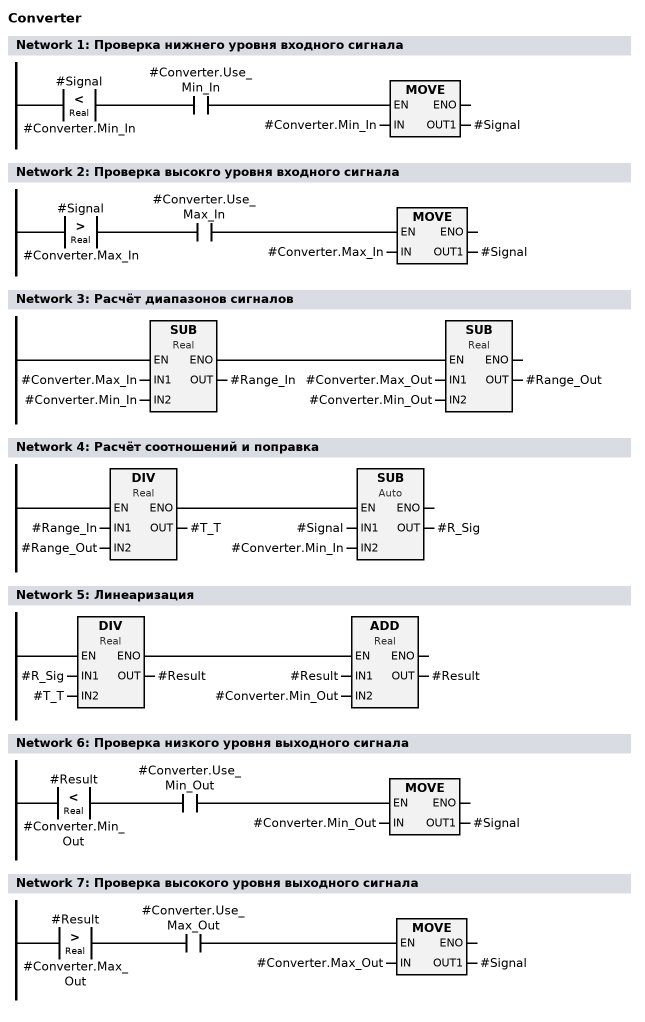
   RUNG wire#powerrail
      { S7_Templates := "SrcType := Real" } LT_Contact(in1 := #Signal, in2 := #Converter.Min_In)
      Contact( #Converter.Use_Min_In )
      Move(in := #Converter.Min_In, out1 => #Signal)
   END_RUNG
   // the same network as SCL:
   IF (#Signal < #Converter.Min_In) AND #Converter.Use_Min_In THEN #Signal := #Converter.Min_In; END_IF;
END_REGION

REGION Network 2: Проверка высокго уровня входного сигнала
   RUNG wire#powerrail
      { S7_Templates := "SrcType := Real" } GT_Contact(in1 := #Signal, in2 := #Converter.Max_In)
      Contact( #Converter.Use_Max_In )
      Move(in := #Converter.Max_In, out1 => #Signal)
   END_RUNG
   // the same network as SCL:
   IF (#Signal > #Converter.Max_In) AND #Converter.Use_Max_In THEN #Signal := #Converter.Max_In; END_IF;
END_REGION

REGION Network 3: Расчёт диапазонов сигналов
   RUNG wire#powerrail
      { S7_Templates := "SrcType := Real"; S7_GenerateENO := "TRUE" } Sub(in1 := #Converter.Max_In, in2 := #Converter.Min_In, out => #Range_In)
      { S7_Templates := "SrcType := Real"; S7_GenerateENO := "TRUE" } Sub(in1 := #Converter.Max_Out, in2 := #Converter.Min_Out, out => #Range_Out)
   END_RUNG
   // the same network as SCL:
   // ENO of a box is taken as its EN; it also drops when the box reports an error
   #Range_In := #Converter.Max_In - #Converter.Min_In;
   #Range_Out := #Converter.Max_Out - #Converter.Min_Out;
END_REGION

REGION Network 4: Расчёт соотношений и поправка
   RUNG wire#powerrail
      { S7_Templates := "SrcType := Real"; S7_GenerateENO := "TRUE" } Div(in1 := #Range_In, in2 := #Range_Out, out => #T_T)
      Sub(in1 := #Signal, in2 := #Converter.Min_In, out => #R_Sig)
   END_RUNG
   // the same network as SCL:
   // ENO of a box is taken as its EN; it also drops when the box reports an error
   #T_T := #Range_In / #Range_Out;
   #R_Sig := #Signal - #Converter.Min_In;
END_REGION

REGION Network 5: Линеаризация
   RUNG wire#powerrail
      { S7_Templates := "SrcType := Real"; S7_GenerateENO := "TRUE" } Div(in1 := #R_Sig, in2 := #T_T, out => #Result)
      { S7_Templates := "SrcType := Real"; S7_GenerateENO := "TRUE" } Add(in1 := #Result, in2 := #Converter.Min_Out, out => #Result)
   END_RUNG
   // the same network as SCL:
   // ENO of a box is taken as its EN; it also drops when the box reports an error
   #Result := #R_Sig / #T_T;
   #Result := #Result + #Converter.Min_Out;
END_REGION

REGION Network 6: Проверка низкого уровня выходного сигнала
   RUNG wire#powerrail
      { S7_Templates := "SrcType := Real" } LT_Contact(in1 := #Result, in2 := #Converter.Min_Out)
      Contact( #Converter.Use_Min_Out )
      Move(in := #Converter.Min_Out, out1 => #Signal)
   END_RUNG
   // the same network as SCL:
   IF (#Result < #Converter.Min_Out) AND #Converter.Use_Min_Out THEN #Signal := #Converter.Min_Out; END_IF;
END_REGION

REGION Network 7: Проверка высокого уровня выходного сигнала
   RUNG wire#powerrail
      { S7_Templates := "SrcType := Real" } GT_Contact(in1 := #Result, in2 := #Converter.Max_Out)
      Contact( #Converter.Use_Max_Out )
      Move(in := #Converter.Max_Out, out1 => #Signal)
   END_RUNG
   // the same network as SCL:
   IF (#Result > #Converter.Max_Out) AND #Converter.Use_Max_Out THEN #Signal := #Converter.Max_Out; END_IF;
END_REGION
END_FUNCTION

FUNCTION "INV" : Void   // FC111, LAD
{ S7_Optimized_Access := 'TRUE' }
VERSION : 0.1
   VAR_INPUT
      S : Bool;   // Сигнал
      I : Bool;   // Инверсия
   END_VAR
   VAR_IN_OUT
      R : Bool;   // Результат
   END_VAR
BEGIN

REGION Network 1: Инверсия сигнала
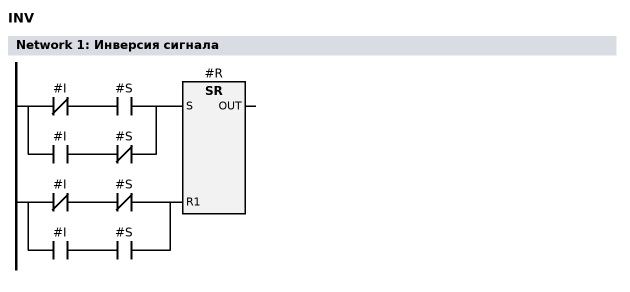
   RUNG wire#powerrail
      I_Contact( #I )
      Contact( #S )
      wire#w1
      S_SR(operand := #R, r1 := wire#w2)
   END_RUNG
   RUNG wire#powerrail
      Contact( #I )
      I_Contact( #S )
   END_RUNG wire#w1
   RUNG wire#powerrail
      I_Contact( #I )
      I_Contact( #S )
   END_RUNG wire#w2
   RUNG wire#powerrail
      Contact( #I )
      Contact( #S )
   END_RUNG wire#w2
   // the same network as SCL:
   IF (NOT #I AND #S) OR (#I AND NOT #S) THEN
       #R := TRUE;   // SR flip-flop
   END_IF;
   IF (NOT #I AND NOT #S) OR (#I AND #S) THEN #R := FALSE; END_IF;
END_REGION
END_FUNCTION

FUNCTION "Mode" : Void   // FC150, LAD
{ S7_Optimized_Access := 'FALSE' }
VERSION : 0.1
   VAR_INPUT
      CMD : Struct   // Основные команды
         Hand : Bool;   // 0 - авто, 1 - ручной / 0 - Авто, 1 - Ручной
         Start_A : Bool;   // Автозапуск / Запуск в авторежиме
         Start_M : Bool;   // Ручной - вперёд / Запуск в ручном режиме
         Force : Bool;   // Принудительный
         Lock : Bool;   // Блокировать / Блокировка
         Local : Bool;   // Локальный
         Service : Bool;   // Сервис
         Safety : Bool;   // Безопасность
         Alarm : Bool;   // Есть авария / Авария
         Reset : Bool;   // Сброс аварий
         Sim : Bool;   // Режим симуляции
      END_STRUCT;
      All_Block : Bool;   // Аварийная блокировка
   END_VAR
   VAR_OUTPUT
      Mode : Int;   // Режим работы
   END_VAR
BEGIN

REGION Network 1: Автоматический режим
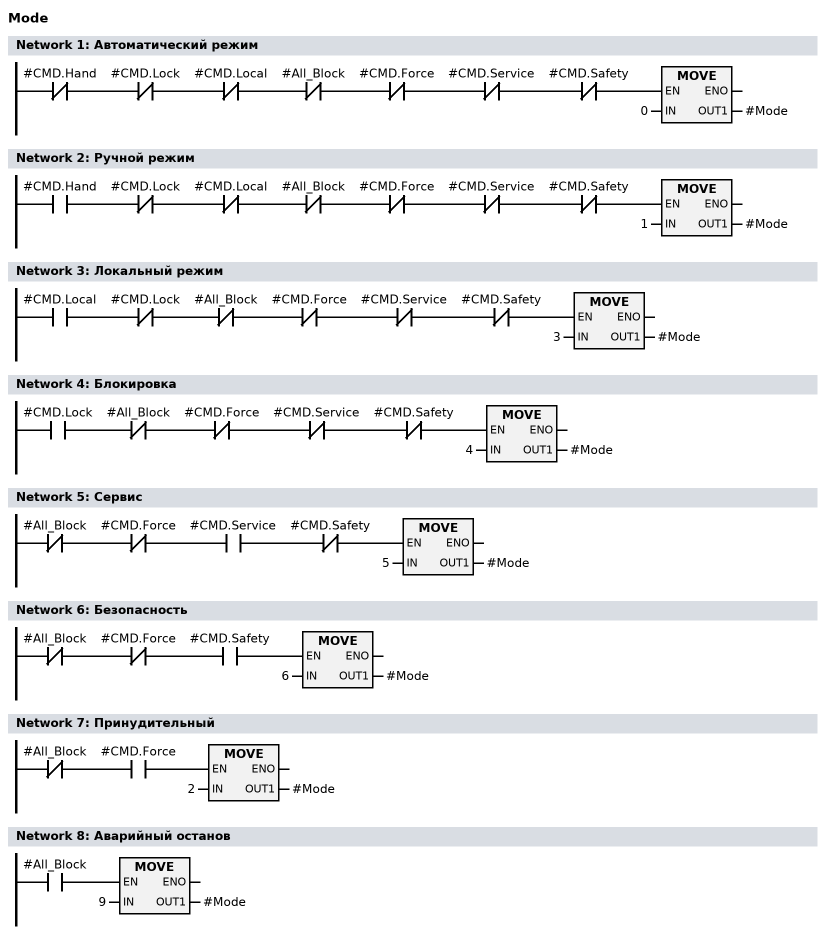
   RUNG wire#powerrail
      I_Contact( #CMD.Hand )
      I_Contact( #CMD.Lock )
      I_Contact( #CMD.Local )
      I_Contact( #All_Block )
      I_Contact( #CMD.Force )
      I_Contact( #CMD.Service )
      I_Contact( #CMD.Safety )
      { S7_GenerateENO := "TRUE" } Move(in := 0, out1 => #Mode)
   END_RUNG
   // the same network as SCL:
   IF NOT #CMD.Hand AND NOT #CMD.Lock AND NOT #CMD.Local AND NOT #All_Block AND NOT #CMD.Force AND NOT #CMD.Service AND NOT #CMD.Safety THEN
       #Mode := 0;
   END_IF;
END_REGION

REGION Network 2: Ручной режим
   RUNG wire#powerrail
      Contact( #CMD.Hand )
      I_Contact( #CMD.Lock )
      I_Contact( #CMD.Local )
      I_Contact( #All_Block )
      I_Contact( #CMD.Force )
      I_Contact( #CMD.Service )
      I_Contact( #CMD.Safety )
      { S7_GenerateENO := "TRUE" } Move(in := 1, out1 => #Mode)
   END_RUNG
   // the same network as SCL:
   IF #CMD.Hand AND NOT #CMD.Lock AND NOT #CMD.Local AND NOT #All_Block AND NOT #CMD.Force AND NOT #CMD.Service AND NOT #CMD.Safety THEN
       #Mode := 1;
   END_IF;
END_REGION

REGION Network 3: Локальный режим
   RUNG wire#powerrail
      Contact( #CMD.Local )
      I_Contact( #CMD.Lock )
      I_Contact( #All_Block )
      I_Contact( #CMD.Force )
      I_Contact( #CMD.Service )
      I_Contact( #CMD.Safety )
      { S7_GenerateENO := "TRUE" } Move(in := 3, out1 => #Mode)
   END_RUNG
   // the same network as SCL:
   IF #CMD.Local AND NOT #CMD.Lock AND NOT #All_Block AND NOT #CMD.Force AND NOT #CMD.Service AND NOT #CMD.Safety THEN
       #Mode := 3;
   END_IF;
END_REGION

REGION Network 4: Блокировка
   RUNG wire#powerrail
      Contact( #CMD.Lock )
      I_Contact( #All_Block )
      I_Contact( #CMD.Force )
      I_Contact( #CMD.Service )
      I_Contact( #CMD.Safety )
      { S7_GenerateENO := "TRUE" } Move(in := 4, out1 => #Mode)
   END_RUNG
   // the same network as SCL:
   IF #CMD.Lock AND NOT #All_Block AND NOT #CMD.Force AND NOT #CMD.Service AND NOT #CMD.Safety THEN
       #Mode := 4;
   END_IF;
END_REGION

REGION Network 5: Сервис
   RUNG wire#powerrail
      I_Contact( #All_Block )
      I_Contact( #CMD.Force )
      Contact( #CMD.Service )
      I_Contact( #CMD.Safety )
      { S7_GenerateENO := "TRUE" } Move(in := 5, out1 => #Mode)
   END_RUNG
   // the same network as SCL:
   IF NOT #All_Block AND NOT #CMD.Force AND #CMD.Service AND NOT #CMD.Safety THEN #Mode := 5; END_IF;
END_REGION

REGION Network 6: Безопасность
   RUNG wire#powerrail
      I_Contact( #All_Block )
      I_Contact( #CMD.Force )
      Contact( #CMD.Safety )
      { S7_GenerateENO := "TRUE" } Move(in := 6, out1 => #Mode)
   END_RUNG
   // the same network as SCL:
   IF NOT #All_Block AND NOT #CMD.Force AND #CMD.Safety THEN #Mode := 6; END_IF;
END_REGION

REGION Network 7: Принудительный
   RUNG wire#powerrail
      I_Contact( #All_Block )
      Contact( #CMD.Force )
      { S7_GenerateENO := "TRUE" } Move(in := 2, out1 => #Mode)
   END_RUNG
   // the same network as SCL:
   IF NOT #All_Block AND #CMD.Force THEN #Mode := 2; END_IF;
END_REGION

REGION Network 8: Аварийный останов
   RUNG wire#powerrail
      Contact( #All_Block )
      { S7_GenerateENO := "TRUE" } Move(in := 9, out1 => #Mode)
   END_RUNG
   // the same network as SCL:
   IF #All_Block THEN #Mode := 9; END_IF;
END_REGION
END_FUNCTION

(* ===== HMI "HMI_RT_1" =====
system functions are stored by id; their names below are inferred from use
connection "HMI_Connection_1": ETHERNET, SMART_S7_1200_OMS

HMI tags "Default tag table"
   "Clock_0.5Hz" : Bool = PLC "Clock_0.5Hz" AT %M0.7, 1 s
   "Mix_1_Clock" : Bool = PLC Mix_1_Clock AT %M10.0, 1 s
   "Mix_2_Clock" : Bool = PLC Mix_2_Clock AT %M10.1, 1 s
   "Mix_3_Clock" : Bool = PLC Mix_3_Clock AT %M10.2, 1 s
   "Logick_DB_Hand" : Bool = PLC Logick_DB.Hand AT %DB1.DBX0.1, 1 s
   "Logick_DB_Start" : Bool = PLC Logick_DB.Start AT %DB1.DBX0.0, 1 s
   "Any_Hand" : Bool = PLC Any_Hand AT %M5.0, 1 s
   "Reset_All" : Bool = PLC Reset_All AT %M3.1, 1 s
   "Logick_DB_T_Probe_SP_S" : Int = PLC Logick_DB.T_Probe.SP_S AT %DB1.DBW60, 1 s
   "Logick_DB_SP_Q" : Real = PLC Logick_DB.SP_Q AT %DB1.DBD2, 1 s
   "Logick_DB_Q" : Real = PLC Logick_DB.Q AT %DB1.DBD6, 1 s
   "Logick_DB_M" : Real = PLC Logick_DB.M AT %DB1.DBD14, 1 s
   "Logick_DB_SP_C" : Real = PLC Logick_DB.SP_C AT %DB1.DBD10, 1 s
   "Any_Alm" : Bool = PLC Any_Alm AT %M6.0, 1 s
   "Logick_DB_M_T" : Real = PLC Logick_DB.M_T AT %DB1.DBD18, 1 s
   "Logick_DB_T_Dos_SP" : Int = PLC Logick_DB.T_Dos.SP AT %DB1.DBW68, 1 s
   "Logick_DB_REQ_Calibration" : Bool = PLC Logick_DB.REQ_Calibration AT %DB1.DBX0.4, 1 s
   "Logick_DB_SP" : Real = PLC Logick_DB.SP AT %DB1.DBD22, 1 s
   "Logick_DB_L_Per_Dos" : Real = PLC Logick_DB.L_Per_Dos AT %DB1.DBD34, 1 s
   "Logick_DB_L_Percent" : Real = PLC Logick_DB.L_Percent AT %DB1.DBD42, 1 s
   "Logick_DB_T_M_SP_M" : Int = PLC Logick_DB.T_M.SP_M AT %DB1.DBW74, 1 s
   "Logick_DB_T_M_1_SP_M" : Int = PLC Logick_DB.T_M_1.SP_M AT %DB1.DBW84, 1 s
   "Logick_DB_T_M_2_SP_M" : Int = PLC Logick_DB.T_M_2.SP_M AT %DB1.DBW94, 1 s
   "Logick_DB_T_M_3_SP_M" : Int = PLC Logick_DB.T_M_3.SP_M AT %DB1.DBW104, 1 s
   "FlowMeter_DB_Full" : Real = PLC FlowMeter_DB.Full AT %DB2.DBD12, 1 s
   "Logick_DB_DD_Stop" : Bool = PLC Logick_DB.DD_Stop AT %DB1.DBX50.2, 1 s
   "Logick_DB_DD_REQ" : Bool = PLC Logick_DB.DD_REQ AT %DB1.DBX50.3, 1 s
   "Logick_DB_T_DD_Stop_SP_M" : Int = PLC Logick_DB.T_DD_Stop.SP_M AT %DB1.DBW134, 1 s
   "Logick_DB_LL_Stop" : Bool = PLC Logick_DB.LL_Stop AT %DB1.DBX50.5, 1 s
   "Logick_DB_HH_Stop" : Bool = PLC Logick_DB.HH_Stop AT %DB1.DBX50.6, 1 s
   "Logick_DB_Level_REQ" : Bool = PLC Logick_DB.Level_REQ AT %DB1.DBX50.7, 1 s
   "Logick_DB_T_Level_Stop_SP_M" : Int = PLC Logick_DB.T_Level_Stop.SP_M AT %DB1.DBW144, 1 s
   "CONFIG_Config_Use_DL" : Bool = PLC CONFIG.Config.Use_DL AT %DB10.DBX0.1, 1 s
   "CONFIG_Config_Use_DD" : Bool = PLC CONFIG.Config.Use_DD AT %DB10.DBX0.0, 1 s
   "CONFIG_Config_Use_Mix_1" : Bool = PLC CONFIG.Config.Use_Mix_1 AT %DB10.DBX0.2, 1 s
   "CONFIG_Config_Use_Mix_2" : Bool = PLC CONFIG.Config.Use_Mix_2 AT %DB10.DBX0.3, 1 s
   "CONFIG_Config_Use_Mix_3" : Bool = PLC CONFIG.Config.Use_Mix_3 AT %DB10.DBX0.4, 1 s
   "DIx_DB_M2_FB_Ready_Inverse" : Bool = PLC DIx_DB.M2_FB_Ready.Inverse AT %DB200.DBX44.3, 1 s
   "DIx_DB_DD_FB_Ready_Inverse" : Bool = PLC DIx_DB.DD_FB_Ready.Inverse AT %DB200.DBX124.3, 1 s
   "Motors_DB_DD_CMD_Sim" : Bool = PLC Motors_DB.DD.CMD.Sim AT %DB204.DBX139.2, 1 s
   "Motors_DB_Vibro_CMD_Sim" : Bool = PLC Motors_DB.Vibro.CMD.Sim AT %DB204.DBX227.2, 1 s
   "Motors_DB_DL_CMD_Sim" : Bool = PLC Motors_DB.DL.CMD.Sim AT %DB204.DBX183.2, 1 s
   "Motors_DB_Mix_1_CMD_Sim" : Bool = PLC Motors_DB.Mix_1.CMD.Sim AT %DB204.DBX7.2, 1 s
   "Motors_DB_Mix_2_CMD_Sim" : Bool = PLC Motors_DB.Mix_2.CMD.Sim AT %DB204.DBX51.2, 1 s
   "Motors_DB_Mix_3_CMD_Sim" : Bool = PLC Motors_DB.Mix_3.CMD.Sim AT %DB204.DBX95.2, 1 s
   "Motors_DB_DD_Status" : Int = PLC Motors_DB.DD.Status AT %DB204.DBW142, 1 s
   "Logick_DB_Alarm" : Word = PLC Logick_DB.Alarm AT %DB1.DBW56, 1 s
   "Motors_DB_Vibro_Status" : Int = PLC Motors_DB.Vibro.Status AT %DB204.DBW230, 1 s
   "Motors_DB_Vibro_Res_h" : DInt = PLC Motors_DB.Vibro.Res_h AT %DB204.DBD256, 1 s
   "Motors_DB_DD_Res_h" : DInt = PLC Motors_DB.DD.Res_h AT %DB204.DBD168, 1 s
   "Any_DB_Level_M" : Int = PLC Any_DB.Level_M AT %DB3.DBW0, 1 s
   "Logick_DB_Level_CMD" : Bool = PLC Logick_DB.Level_CMD AT %DB1.DBX51.0, 1 s
   "Any_DB_Flow_M" : Int = PLC Any_DB.Flow_M AT %DB3.DBW4, 1 s
   "Logick_DB_DD_CMD" : Bool = PLC Logick_DB.DD_CMD AT %DB1.DBX50.4, 1 s
   "Any_DB_DD_View" : Bool = PLC Any_DB.DD_View AT %DB3.DBX8.0, 1 s
   "Any_DB_Level_View" : Bool = PLC Any_DB.Level_View AT %DB3.DBX8.1, 1 s
   "AIx_DB_Level_Alarms_LL" : Bool = PLC AIx_DB.Level.Alarms.LL AT %DB202.DBX276.5, 1 s
   "AIx_DB_Level_Alarms_HH" : Bool = PLC AIx_DB.Level.Alarms.HH AT %DB202.DBX276.2, 1 s

HMI tags "HMI"
   "settings" : Int, internal

HMI tags "xDI"
   "DIx_DB_Vibro_FB_Ready_Signal" : Bool = PLC DIx_DB.Vibro_FB_Ready.Signal AT %DB200.DBX182.0, 1 s
   "DIx_DB_Transporter_Signal" : Bool = PLC DIx_DB.Transporter.Signal AT %DB200.DBX202.0, 1 s
   "DIx_DB_M3_FB_Run_Signal" : Bool = PLC DIx_DB.M3_FB_Run.Signal AT %DB200.DBX102.0, 1 s
   "DIx_DB_M3_FB_Ready_Signal" : Bool = PLC DIx_DB.M3_FB_Ready.Signal AT %DB200.DBX82.0, 1 s
   "DIx_DB_M2_FB_Run_Signal" : Bool = PLC DIx_DB.M2_FB_Run.Signal AT %DB200.DBX62.0, 1 s
   "DIx_DB_M2_FB_Ready_Signal" : Bool = PLC DIx_DB.M2_FB_Ready.Signal AT %DB200.DBX42.0, 1 s
   "DIx_DB_M1_FB_Run_Signal" : Bool = PLC DIx_DB.M1_FB_Run.Signal AT %DB200.DBX22.0, 1 s
   "DIx_DB_M1_FB_Ready_Signal" : Bool = PLC DIx_DB.M1_FB_Ready.Signal AT %DB200.DBX2.0, 1 s
   "DIx_DB_Flow_Signal" : Bool = PLC DIx_DB.Dry_Run.Signal AT %DB200.DBX242.0, 1 s
   "DIx_DB_Dos_FB_Run_Signal" : Bool = PLC DIx_DB.Dos_FB_Run.Signal AT %DB200.DBX142.0, 1 s
   "DIx_DB_DL_FB_Ready_Signal" : Bool = PLC DIx_DB.DL_FB_Ready.Signal AT %DB200.DBX222.0, 1 s
   "DIx_DB_DD_LLS_Signal" : Bool = PLC DIx_DB.DD_LLS.Signal AT %DB200.DBX162.0, 1 s
   "DIx_DB_DD_FB_Ready_Signal" : Bool = PLC DIx_DB.DD_FB_Ready.Signal AT %DB200.DBX122.0, 1 s
   "DIx_DB_AllBlock_Signal" : Bool = PLC DIx_DB.AllBlock.Signal AT %DB200.DBX262.0, 1 s
   "DIx_DB_M1_FB_Ready_Input" : Bool = PLC DIx_DB.M1_FB_Ready.Input AT %DB200.DBX0.0, 1 s
   "DIx_DB_M1_FB_Ready_Hand" : Bool = PLC DIx_DB.M1_FB_Ready.Hand AT %DB200.DBX4.0, 1 s
   "DIx_DB_M1_FB_Ready_Start_M" : Bool = PLC DIx_DB.M1_FB_Ready.Start_M AT %DB200.DBX4.1, 1 s
   "DIx_DB_M1_FB_Ready_Inverse" : Bool = PLC DIx_DB.M1_FB_Ready.Inverse AT %DB200.DBX4.3, 1 s
   "DIx_DB_M1_FB_Ready_Filter_On_SP" : Int = PLC DIx_DB.M1_FB_Ready.Filter_On.SP AT %DB200.DBW6, 1 s
   "DIx_DB_M1_FB_Ready_Filter_Off_SP" : Int = PLC DIx_DB.M1_FB_Ready.Filter_Off.SP AT %DB200.DBW12, 1 s
   "DIx_DB_M1_FB_Run_Input" : Bool = PLC DIx_DB.M1_FB_Run.Input AT %DB200.DBX20.0, 1 s
   "DIx_DB_M1_FB_Run_Hand" : Bool = PLC DIx_DB.M1_FB_Run.Hand AT %DB200.DBX24.0, 1 s
   "DIx_DB_M1_FB_Run_Start_M" : Bool = PLC DIx_DB.M1_FB_Run.Start_M AT %DB200.DBX24.1, 1 s
   "DIx_DB_M1_FB_Run_Inverse" : Bool = PLC DIx_DB.M1_FB_Run.Inverse AT %DB200.DBX24.3, 1 s
   "DIx_DB_M1_FB_Run_Filter_On_SP" : Int = PLC DIx_DB.M1_FB_Run.Filter_On.SP AT %DB200.DBW26, 1 s
   "DIx_DB_M1_FB_Run_Filter_Off_SP" : Int = PLC DIx_DB.M1_FB_Run.Filter_Off.SP AT %DB200.DBW32, 1 s
   "DIx_DB_M2_FB_Ready_Filter_Off_SP" : Int = PLC DIx_DB.M2_FB_Ready.Filter_Off.SP AT %DB200.DBW52, 1 s
   "DIx_DB_M2_FB_Ready_Filter_On_SP" : Int = PLC DIx_DB.M2_FB_Ready.Filter_On.SP AT %DB200.DBW46, 1 s
   "DIx_DB_M2_FB_Ready_Hand" : Bool = PLC DIx_DB.M2_FB_Ready.Hand AT %DB200.DBX44.0, 1 s
   "DIx_DB_M2_FB_Ready_Start_M" : Bool = PLC DIx_DB.M2_FB_Ready.Start_M AT %DB200.DBX44.1, 1 s
   "DIx_DB_M2_FB_Ready_Input" : Bool = PLC DIx_DB.M2_FB_Ready.Input AT %DB200.DBX40.0, 1 s
   "DIx_DB_M2_FB_Run_Input" : Bool = PLC DIx_DB.M2_FB_Run.Input AT %DB200.DBX60.0, 1 s
   "DIx_DB_M2_FB_Run_Hand" : Bool = PLC DIx_DB.M2_FB_Run.Hand AT %DB200.DBX64.0, 1 s
   "DIx_DB_M2_FB_Run_Start_M" : Bool = PLC DIx_DB.M2_FB_Run.Start_M AT %DB200.DBX64.1, 1 s
   "DIx_DB_M2_FB_Run_Inverse" : Bool = PLC DIx_DB.M2_FB_Run.Inverse AT %DB200.DBX64.3, 1 s
   "DIx_DB_M2_FB_Run_Filter_On_SP" : Int = PLC DIx_DB.M2_FB_Run.Filter_On.SP AT %DB200.DBW66, 1 s
   "DIx_DB_M2_FB_Run_Filter_Off_SP" : Int = PLC DIx_DB.M2_FB_Run.Filter_Off.SP AT %DB200.DBW72, 1 s
   "DIx_DB_M3_FB_Ready_Input" : Bool = PLC DIx_DB.M3_FB_Ready.Input AT %DB200.DBX80.0, 1 s
   "DIx_DB_M3_FB_Ready_Hand" : Bool = PLC DIx_DB.M3_FB_Ready.Hand AT %DB200.DBX84.0, 1 s
   "DIx_DB_M3_FB_Ready_Start_M" : Bool = PLC DIx_DB.M3_FB_Ready.Start_M AT %DB200.DBX84.1, 1 s
   "DIx_DB_M3_FB_Ready_Inverse" : Bool = PLC DIx_DB.M3_FB_Ready.Inverse AT %DB200.DBX84.3, 1 s
   "DIx_DB_M3_FB_Ready_Filter_On_SP" : Int = PLC DIx_DB.M3_FB_Ready.Filter_On.SP AT %DB200.DBW86, 1 s
   "DIx_DB_M3_FB_Ready_Filter_Off_SP" : Int = PLC DIx_DB.M3_FB_Ready.Filter_Off.SP AT %DB200.DBW92, 1 s
   "DIx_DB_M3_FB_Run_Input" : Bool = PLC DIx_DB.M3_FB_Run.Input AT %DB200.DBX100.0, 1 s
   "DIx_DB_M3_FB_Run_Hand" : Bool = PLC DIx_DB.M3_FB_Run.Hand AT %DB200.DBX104.0, 1 s
   "DIx_DB_M3_FB_Run_Start_M" : Bool = PLC DIx_DB.M3_FB_Run.Start_M AT %DB200.DBX104.1, 1 s
   "DIx_DB_M3_FB_Run_Inverse" : Bool = PLC DIx_DB.M3_FB_Run.Inverse AT %DB200.DBX104.3, 1 s
   "DIx_DB_M3_FB_Run_Filter_On_SP" : Int = PLC DIx_DB.M3_FB_Run.Filter_On.SP AT %DB200.DBW106, 1 s
   "DIx_DB_M3_FB_Run_Filter_Off_SP" : Int = PLC DIx_DB.M3_FB_Run.Filter_Off.SP AT %DB200.DBW112, 1 s
   "DIx_DB_DD_FB_Ready_Input" : Bool = PLC DIx_DB.DD_FB_Ready.Input AT %DB200.DBX120.0, 1 s
   "DIx_DB_DD_FB_Ready_Hand" : Bool = PLC DIx_DB.DD_FB_Ready.Hand AT %DB200.DBX124.0, 1 s
   "DIx_DB_DD_FB_Ready_Start_M" : Bool = PLC DIx_DB.DD_FB_Ready.Start_M AT %DB200.DBX124.1, 1 s
   "DIx_DB_DD_FB_Ready_Filter_On_SP" : Int = PLC DIx_DB.DD_FB_Ready.Filter_On.SP AT %DB200.DBW126, 1 s
   "DIx_DB_DD_FB_Ready_Filter_Off_SP" : Int = PLC DIx_DB.DD_FB_Ready.Filter_Off.SP AT %DB200.DBW132, 1 s
   "DIx_DB_Dos_FB_Run_Input" : Bool = PLC DIx_DB.Dos_FB_Run.Input AT %DB200.DBX140.0, 1 s
   "DIx_DB_Dos_FB_Run_Hand" : Bool = PLC DIx_DB.Dos_FB_Run.Hand AT %DB200.DBX144.0, 1 s
   "DIx_DB_Dos_FB_Run_Start_M" : Bool = PLC DIx_DB.Dos_FB_Run.Start_M AT %DB200.DBX144.1, 1 s
   "DIx_DB_Dos_FB_Run_Inverse" : Bool = PLC DIx_DB.Dos_FB_Run.Inverse AT %DB200.DBX144.3, 1 s
   "DIx_DB_Dos_FB_Run_Filter_On_SP" : Int = PLC DIx_DB.Dos_FB_Run.Filter_On.SP AT %DB200.DBW146, 1 s
   "DIx_DB_Dos_FB_Run_Filter_Off_SP" : Int = PLC DIx_DB.Dos_FB_Run.Filter_Off.SP AT %DB200.DBW152, 1 s
   "DIx_DB_DD_LLS_Input" : Bool = PLC DIx_DB.DD_LLS.Input AT %DB200.DBX160.0, 1 s
   "DIx_DB_DD_LLS_Hand" : Bool = PLC DIx_DB.DD_LLS.Hand AT %DB200.DBX164.0, 1 s
   "DIx_DB_DD_LLS_Start_M" : Bool = PLC DIx_DB.DD_LLS.Start_M AT %DB200.DBX164.1, 1 s
   "DIx_DB_DD_LLS_Inverse" : Bool = PLC DIx_DB.DD_LLS.Inverse AT %DB200.DBX164.3, 1 s
   "DIx_DB_DD_LLS_Filter_On_SP" : Int = PLC DIx_DB.DD_LLS.Filter_On.SP AT %DB200.DBW166, 1 s
   "DIx_DB_DD_LLS_Filter_Off_SP" : Int = PLC DIx_DB.DD_LLS.Filter_Off.SP AT %DB200.DBW172, 1 s
   "DIx_DB_Vibro_FB_Ready_Input" : Bool = PLC DIx_DB.Vibro_FB_Ready.Input AT %DB200.DBX180.0, 1 s
   "DIx_DB_Vibro_FB_Ready_Hand" : Bool = PLC DIx_DB.Vibro_FB_Ready.Hand AT %DB200.DBX184.0, 1 s
   "DIx_DB_Vibro_FB_Ready_Start_M" : Bool = PLC DIx_DB.Vibro_FB_Ready.Start_M AT %DB200.DBX184.1, 1 s
   "DIx_DB_Vibro_FB_Ready_Inverse" : Bool = PLC DIx_DB.Vibro_FB_Ready.Inverse AT %DB200.DBX184.3, 1 s
   "DIx_DB_Vibro_FB_Ready_Filter_On_SP" : Int = PLC DIx_DB.Vibro_FB_Ready.Filter_On.SP AT %DB200.DBW186, 1 s
   "DIx_DB_Vibro_FB_Ready_Filter_Off_SP" : Int = PLC DIx_DB.Vibro_FB_Ready.Filter_Off.SP AT %DB200.DBW192, 1 s
   "DIx_DB_Transporter_Input" : Bool = PLC DIx_DB.Transporter.Input AT %DB200.DBX200.0, 1 s
   "DIx_DB_Transporter_Hand" : Bool = PLC DIx_DB.Transporter.Hand AT %DB200.DBX204.0, 1 s
   "DIx_DB_Transporter_Start_M" : Bool = PLC DIx_DB.Transporter.Start_M AT %DB200.DBX204.1, 1 s
   "DIx_DB_Transporter_Inverse" : Bool = PLC DIx_DB.Transporter.Inverse AT %DB200.DBX204.3, 1 s
   "DIx_DB_Transporter_Filter_On_SP" : Int = PLC DIx_DB.Transporter.Filter_On.SP AT %DB200.DBW206, 1 s
   "DIx_DB_Transporter_Filter_Off_SP" : Int = PLC DIx_DB.Transporter.Filter_Off.SP AT %DB200.DBW212, 1 s
   "DIx_DB_DL_FB_Ready_Input" : Bool = PLC DIx_DB.DL_FB_Ready.Input AT %DB200.DBX220.0, 1 s
   "DIx_DB_DL_FB_Ready_Hand" : Bool = PLC DIx_DB.DL_FB_Ready.Hand AT %DB200.DBX224.0, 1 s
   "DIx_DB_DL_FB_Ready_Start_M" : Bool = PLC DIx_DB.DL_FB_Ready.Start_M AT %DB200.DBX224.1, 1 s
   "DIx_DB_DL_FB_Ready_Inverse" : Bool = PLC DIx_DB.DL_FB_Ready.Inverse AT %DB200.DBX224.3, 1 s
   "DIx_DB_DL_FB_Ready_Filter_On_SP" : Int = PLC DIx_DB.DL_FB_Ready.Filter_On.SP AT %DB200.DBW226, 1 s
   "DIx_DB_DL_FB_Ready_Filter_Off_SP" : Int = PLC DIx_DB.DL_FB_Ready.Filter_Off.SP AT %DB200.DBW232, 1 s
   "DIx_DB_Flow_Input" : Bool = PLC DIx_DB.Dry_Run.Input AT %DB200.DBX240.0, 1 s
   "DIx_DB_Flow_Hand" : Bool = PLC DIx_DB.Dry_Run.Hand AT %DB200.DBX244.0, 1 s
   "DIx_DB_Flow_Start_M" : Bool = PLC DIx_DB.Dry_Run.Start_M AT %DB200.DBX244.1, 1 s
   "DIx_DB_Flow_Inverse" : Bool = PLC DIx_DB.Dry_Run.Inverse AT %DB200.DBX244.3, 1 s
   "DIx_DB_Flow_Filter_On_SP" : Int = PLC DIx_DB.Dry_Run.Filter_On.SP AT %DB200.DBW246, 1 s
   "DIx_DB_Flow_Filter_Off_SP" : Int = PLC DIx_DB.Dry_Run.Filter_Off.SP AT %DB200.DBW252, 1 s
   "DIx_DB_AllBlock_Filter_Off_SP" : Int = PLC DIx_DB.AllBlock.Filter_Off.SP AT %DB200.DBW272, 1 s
   "DIx_DB_AllBlock_Filter_On_SP" : Int = PLC DIx_DB.AllBlock.Filter_On.SP AT %DB200.DBW266, 1 s
   "DIx_DB_AllBlock_Inverse" : Bool = PLC DIx_DB.AllBlock.Inverse AT %DB200.DBX264.3, 1 s
   "DIx_DB_AllBlock_Start_M" : Bool = PLC DIx_DB.AllBlock.Start_M AT %DB200.DBX264.1, 1 s
   "DIx_DB_AllBlock_Hand" : Bool = PLC DIx_DB.AllBlock.Hand AT %DB200.DBX264.0, 1 s
   "DIx_DB_AllBlock_Input" : Bool = PLC DIx_DB.AllBlock.Input AT %DB200.DBX260.0, 1 s

HMI tags "xDO"
   "DOx_DB_Vibro_CMD_Q" : Bool = PLC DOx_DB.Vibro_CMD.Q AT %DB201.DBX40.2, 1 s
   "DOx_DB_M3_CMD_Q" : Bool = PLC DOx_DB.M3_CMD.Q AT %DB201.DBX20.2, 1 s
   "DOx_DB_M2_CMD_Q" : Bool = PLC DOx_DB.M2_CMD.Q AT %DB201.DBX10.2, 1 s
   "DOx_DB_M1_CMD_Q" : Bool = PLC DOx_DB.M1_CMD.Q AT %DB201.DBX0.2, 1 s
   "DOx_DB_LED_Empty_Q" : Bool = PLC DOx_DB.LED_Empty.Q AT %DB201.DBX90.2, 1 s
   "DOx_DB_LED_Dry_Run_Q" : Bool = PLC DOx_DB.LED_Dry_Run.Q AT %DB201.DBX70.2, 1 s
   "DOx_DB_LED_Alarm_Q" : Bool = PLC DOx_DB.LED_Alarm.Q AT %DB201.DBX80.2, 1 s
   "DOx_DB_KC1_CMD_Q" : Bool = PLC DOx_DB.KC1_CMD.Q AT %DB201.DBX60.2, 1 s
   "DOx_DB_DL_CMD_Q" : Bool = PLC DOx_DB.DL_CMD.Q AT %DB201.DBX50.2, 1 s
   "DOx_DB_DD_CMD_Q" : Bool = PLC DOx_DB.DD_CMD.Q AT %DB201.DBX30.2, 1 s
   "DOx_DB_M1_CMD_Start_A" : Bool = PLC DOx_DB.M1_CMD.Start_A AT %DB201.DBX0.0, 1 s
   "DOx_DB_M1_CMD_Hand" : Bool = PLC DOx_DB.M1_CMD.Hand AT %DB201.DBX2.0, 1 s
   "DOx_DB_M1_CMD_Start_M" : Bool = PLC DOx_DB.M1_CMD.Start_M AT %DB201.DBX2.1, 1 s
   "DOx_DB_M1_CMD_Simulation" : Bool = PLC DOx_DB.M1_CMD.Simulation AT %DB201.DBX2.2, 1 s
   "DOx_DB_M1_CMD_Inverse" : Bool = PLC DOx_DB.M1_CMD.Inverse AT %DB201.DBX2.3, 1 s
   "DOx_DB_M2_CMD_Start_A" : Bool = PLC DOx_DB.M2_CMD.Start_A AT %DB201.DBX10.0, 1 s
   "DOx_DB_M2_CMD_Hand" : Bool = PLC DOx_DB.M2_CMD.Hand AT %DB201.DBX12.0, 1 s
   "DOx_DB_M2_CMD_Start_M" : Bool = PLC DOx_DB.M2_CMD.Start_M AT %DB201.DBX12.1, 1 s
   "DOx_DB_M2_CMD_Simulation" : Bool = PLC DOx_DB.M2_CMD.Simulation AT %DB201.DBX12.2, 1 s
   "DOx_DB_M2_CMD_Inverse" : Bool = PLC DOx_DB.M2_CMD.Inverse AT %DB201.DBX12.3, 1 s
   "DOx_DB_M3_CMD_Start_A" : Bool = PLC DOx_DB.M3_CMD.Start_A AT %DB201.DBX20.0, 1 s
   "DOx_DB_M3_CMD_Hand" : Bool = PLC DOx_DB.M3_CMD.Hand AT %DB201.DBX22.0, 1 s
   "DOx_DB_M3_CMD_Start_M" : Bool = PLC DOx_DB.M3_CMD.Start_M AT %DB201.DBX22.1, 1 s
   "DOx_DB_M3_CMD_Simulation" : Bool = PLC DOx_DB.M3_CMD.Simulation AT %DB201.DBX22.2, 1 s
   "DOx_DB_M3_CMD_Inverse" : Bool = PLC DOx_DB.M3_CMD.Inverse AT %DB201.DBX22.3, 1 s
   "DOx_DB_DD_CMD_Start_A" : Bool = PLC DOx_DB.DD_CMD.Start_A AT %DB201.DBX30.0, 1 s
   "DOx_DB_DD_CMD_Hand" : Bool = PLC DOx_DB.DD_CMD.Hand AT %DB201.DBX32.0, 1 s
   "DOx_DB_DD_CMD_Start_M" : Bool = PLC DOx_DB.DD_CMD.Start_M AT %DB201.DBX32.1, 1 s
   "DOx_DB_DD_CMD_Simulation" : Bool = PLC DOx_DB.DD_CMD.Simulation AT %DB201.DBX32.2, 1 s
   "DOx_DB_DD_CMD_Inverse" : Bool = PLC DOx_DB.DD_CMD.Inverse AT %DB201.DBX32.3, 1 s
   "DOx_DB_Vibro_CMD_Start_A" : Bool = PLC DOx_DB.Vibro_CMD.Start_A AT %DB201.DBX40.0, 1 s
   "DOx_DB_Vibro_CMD_Hand" : Bool = PLC DOx_DB.Vibro_CMD.Hand AT %DB201.DBX42.0, 1 s
   "DOx_DB_Vibro_CMD_Start_M" : Bool = PLC DOx_DB.Vibro_CMD.Start_M AT %DB201.DBX42.1, 1 s
   "DOx_DB_Vibro_CMD_Simulation" : Bool = PLC DOx_DB.Vibro_CMD.Simulation AT %DB201.DBX42.2, 1 s
   "DOx_DB_Vibro_CMD_Inverse" : Bool = PLC DOx_DB.Vibro_CMD.Inverse AT %DB201.DBX42.3, 1 s
   "DOx_DB_DL_CMD_Start_A" : Bool = PLC DOx_DB.DL_CMD.Start_A AT %DB201.DBX50.0, 1 s
   "DOx_DB_DL_CMD_Hand" : Bool = PLC DOx_DB.DL_CMD.Hand AT %DB201.DBX52.0, 1 s
   "DOx_DB_DL_CMD_Start_M" : Bool = PLC DOx_DB.DL_CMD.Start_M AT %DB201.DBX52.1, 1 s
   "DOx_DB_DL_CMD_Simulation" : Bool = PLC DOx_DB.DL_CMD.Simulation AT %DB201.DBX52.2, 1 s
   "DOx_DB_DL_CMD_Inverse" : Bool = PLC DOx_DB.DL_CMD.Inverse AT %DB201.DBX52.3, 1 s
   "DOx_DB_KC1_CMD_Start_A" : Bool = PLC DOx_DB.KC1_CMD.Start_A AT %DB201.DBX60.0, 1 s
   "DOx_DB_KC1_CMD_Hand" : Bool = PLC DOx_DB.KC1_CMD.Hand AT %DB201.DBX62.0, 1 s
   "DOx_DB_KC1_CMD_Start_M" : Bool = PLC DOx_DB.KC1_CMD.Start_M AT %DB201.DBX62.1, 1 s
   "DOx_DB_KC1_CMD_Simulation" : Bool = PLC DOx_DB.KC1_CMD.Simulation AT %DB201.DBX62.2, 1 s
   "DOx_DB_KC1_CMD_Inverse" : Bool = PLC DOx_DB.KC1_CMD.Inverse AT %DB201.DBX62.3, 1 s
   "DOx_DB_LED_Dry_Run_Start_A" : Bool = PLC DOx_DB.LED_Dry_Run.Start_A AT %DB201.DBX70.0, 1 s
   "DOx_DB_LED_Dry_Run_Hand" : Bool = PLC DOx_DB.LED_Dry_Run.Hand AT %DB201.DBX72.0, 1 s
   "DOx_DB_LED_Dry_Run_Start_M" : Bool = PLC DOx_DB.LED_Dry_Run.Start_M AT %DB201.DBX72.1, 1 s
   "DOx_DB_LED_Dry_Run_Simulation" : Bool = PLC DOx_DB.LED_Dry_Run.Simulation AT %DB201.DBX72.2, 1 s
   "DOx_DB_LED_Dry_Run_Inverse" : Bool = PLC DOx_DB.LED_Dry_Run.Inverse AT %DB201.DBX72.3, 1 s
   "DOx_DB_LED_Alarm_Start_A" : Bool = PLC DOx_DB.LED_Alarm.Start_A AT %DB201.DBX80.0, 1 s
   "DOx_DB_LED_Alarm_Hand" : Bool = PLC DOx_DB.LED_Alarm.Hand AT %DB201.DBX82.0, 1 s
   "DOx_DB_LED_Alarm_Start_M" : Bool = PLC DOx_DB.LED_Alarm.Start_M AT %DB201.DBX82.1, 1 s
   "DOx_DB_LED_Alarm_Simulation" : Bool = PLC DOx_DB.LED_Alarm.Simulation AT %DB201.DBX82.2, 1 s
   "DOx_DB_LED_Alarm_Inverse" : Bool = PLC DOx_DB.LED_Alarm.Inverse AT %DB201.DBX82.3, 1 s
   "DOx_DB_LED_Empty_Start_A" : Bool = PLC DOx_DB.LED_Empty.Start_A AT %DB201.DBX90.0, 1 s
   "DOx_DB_LED_Empty_Hand" : Bool = PLC DOx_DB.LED_Empty.Hand AT %DB201.DBX92.0, 1 s
   "DOx_DB_LED_Empty_Start_M" : Bool = PLC DOx_DB.LED_Empty.Start_M AT %DB201.DBX92.1, 1 s
   "DOx_DB_LED_Empty_Simulation" : Bool = PLC DOx_DB.LED_Empty.Simulation AT %DB201.DBX92.2, 1 s
   "DOx_DB_LED_Empty_Inverse" : Bool = PLC DOx_DB.LED_Empty.Inverse AT %DB201.DBX92.3, 1 s
